   "86_Times_STEP_MAX_TIME_STP_010(1)" : Time = PLC "86_Times".STEP_MAX_TIME_STP_010 AT %DB1.DBW0, 1 s
   "86_Times_STEP_MAX_TIME_STP_020(1)" : Time = PLC "86_Times".STEP_MAX_TIME_STP_020 AT %DB1.DBW0, 1 s
   "86_Times_STEP_MAX_TIME_STP_030(1)" : Time = PLC "86_Times".STEP_MAX_TIME_STP_030 AT %DB1.DBW0, 1 s
   "86_Times_STEP_MAX_TIME_STP_040(1)" : Time = PLC "86_Times".STEP_MAX_TIME_STP_040 AT %DB1.DBW0, 1 s
   "86_Times_STEP_MAX_TIME_STP_050(1)" : Time = PLC "86_Times".STEP_MAX_TIME_STP_050 AT %DB1.DBW0, 1 s
   "86_Times_STEP_MAX_TIME_STP_060(1)" : Time = PLC "86_Times".STEP_MAX_TIME_STP_060 AT %DB1.DBW0, 1 s
   "86_Times_STEP_MAX_TIME_STP_070(1)" : Time = PLC "86_Times".STEP_MAX_TIME_STP_070 AT %DB1.DBW0, 1 s
   "86_Times_STEP_MAX_TIME_STP_080(1)" : Time = PLC "86_Times".STEP_MAX_TIME_STP_080 AT %DB1.DBW0, 1 s
   "86_Times_STEP_MAX_TIME_STP_090(1)" : Time = PLC "86_Times".STEP_MAX_TIME_STP_090 AT %DB1.DBW0, 1 s
   "86_Times_STEP_MAX_TIME_STP_100(1)" : Time = PLC "86_Times".STEP_MAX_TIME_STP_100 AT %DB1.DBW0, 1 s
   "86_Times_STEP_MAX_TIME_STP_110(1)" : Time = PLC "86_Times".STEP_MAX_TIME_STP_110 AT %DB1.DBW0, 1 s
   "86_Times_STEP_MAX_TIME_STP_120(1)" : Time = PLC "86_Times".STEP_MAX_TIME_STP_120 AT %DB1.DBW0, 1 s
   "86_Times_STEP_MAX_TIME_STP_130(1)" : Time = PLC "86_Times".STEP_MAX_TIME_STP_130 AT %DB1.DBW0, 1 s
   "86_Times_STEP_MAX_TIME_STP_140(1)" : Time = PLC "86_Times".STEP_MAX_TIME_STP_140 AT %DB1.DBW0, 1 s
   "86_Times_STEP_MAX_TIME_STP_150(1)" : Time = PLC "86_Times".STEP_MAX_TIME_STP_150 AT %DB1.DBW0, 1 s
   "86_Times_STEP_MAX_TIME_STP_160(1)" : Time = PLC "86_Times".STEP_MAX_TIME_STP_160 AT %DB1.DBW0, 1 s
   "86_Times_STEP_MAX_TIME_STP_170(1)" : Time = PLC "86_Times".STEP_MAX_TIME_STP_170 AT %DB1.DBW0, 1 s
   "86_Times_STEP_MAX_TIME_STP_180(1)" : Time = PLC "86_Times".STEP_MAX_TIME_STP_180 AT %DB1.DBW0, 1 s
   "86_Times_STEP_MAX_TIME_STP_190(1)" : Time = PLC "86_Times".STEP_MAX_TIME_STP_190 AT %DB1.DBW0, 1 s
   "86_Times_STEP_MAX_TIME_STP_200(1)" : Time = PLC "86_Times".STEP_MAX_TIME_STP_200 AT %DB1.DBW0, 1 s
   "86_Times_STEP_MAX_TIME_STP_210(1)" : Time = PLC "86_Times".STEP_MAX_TIME_STP_210 AT %DB1.DBW0, 1 s
   "86_Times_STEP_MAX_TIME_STP_220(1)" : Time = PLC "86_Times".STEP_MAX_TIME_STP_220 AT %DB1.DBW0, 1 s
   "86_Times_STEP_MAX_TIME_STP_230(1)" : Time = PLC "86_Times".STEP_MAX_TIME_STP_230 AT %DB1.DBW0, 1 s
   "86_Times_STEP_MAX_TIME_STP_240(1)" : Time = PLC "86_Times".STEP_MAX_TIME_STP_240 AT %DB1.DBW0, 1 s
   "86_Times_STEP_MAX_TIME_STP_250(1)" : Time = PLC "86_Times".STEP_MAX_TIME_STP_250 AT %DB1.DBW0, 1 s
   "86_Times_STEP_MAX_TIME_STP_260(1)" : Time = PLC "86_Times".STEP_MAX_TIME_STP_260 AT %DB1.DBW0, 1 s
   "86_Times_STEP_MAX_TIME_STP_270(1)" : Time = PLC "86_Times".STEP_MAX_TIME_STP_270 AT %DB1.DBW0, 1 s
   "86_Times_STEP_MAX_TIME_STP_280(1)" : Time = PLC "86_Times".STEP_MAX_TIME_STP_280 AT %DB1.DBW0, 1 s
   "86_Times_STEP_MAX_TIME_STP_290(1)" : Time = PLC "86_Times".STEP_MAX_TIME_STP_290 AT %DB1.DBW0, 1 s
   "86_Times_STEP_MAX_TIME_STP_300(1)" : Time = PLC "86_Times".STEP_MAX_TIME_STP_300 AT %DB1.DBW0, 1 s
   "86_Times_STEP_MAX_TIME_STP_310(1)" : Time = PLC "86_Times".STEP_MAX_TIME_STP_310 AT %DB1.DBW0, 1 s
   "86_Times_STEP_MAX_TIME_STP_320(1)" : Time = PLC "86_Times".STEP_MAX_TIME_STP_320 AT %DB1.DBW0, 1 s
   "86_Times_STEP_MAX_TIME_STP_330(1)" : Time = PLC "86_Times".STEP_MAX_TIME_STP_330 AT %DB1.DBW0, 1 s
   "86_Times_STEP_MAX_TIME_STP_340(1)" : Time = PLC "86_Times".STEP_MAX_TIME_STP_340 AT %DB1.DBW0, 1 s
   "86_Times_STEP_MAX_TIME_STP_350(1)" : Time = PLC Alarms_Acknowledge.IGG_ALARM_ACKNLG_2 AT %DB1.DBW0, 1 s
   "86_Times_STEP_MAX_TIME_STP_360(1)" : Time = PLC "86_Times".STEP_MAX_TIME_STP_360 AT %DB1.DBW0, 1 s
   "86_Times_STEP_MAX_TIME_STP_370(1)" : Time = PLC "86_Times".STEP_MAX_TIME_STP_370 AT %DB1.DBW0, 1 s
   "86_Times_STEP_MAX_TIME_STP_380(1)" : Time = PLC "86_Times".STEP_MAX_TIME_STP_380 AT %DB1.DBW0, 1 s
   "86_Times_STEP_MAX_TIME_STP_390(1)" : Time = PLC "86_Times".STEP_MAX_TIME_STP_390 AT %DB1.DBW0, 1 s
   "86_Times_STEP_MAX_TIME_STP_400(1)" : Time = PLC "86_Times".STEP_MAX_TIME_STP_400 AT %DB1.DBW0, 1 s
   "86_Times_STEP_MAX_TIME_STP_410(1)" : Time = PLC "86_Times".STEP_MAX_TIME_STP_410 AT %DB1.DBW0, 1 s
   "86_Times_STEP_MAX_TIME_STP_420(1)" : Time = PLC "86_Times".STEP_MAX_TIME_STP_420 AT %DB1.DBW0, 1 s
   "86_Times_STEP_MAX_TIME_STP_430(1)" : Time = PLC "86_Times".STEP_MAX_TIME_STP_430 AT %DB1.DBW0, 1 s
   "86_Times_STEP_MAX_TIME_STP_440(1)" : Time = PLC "86_Times".STEP_MAX_TIME_STP_440 AT %DB1.DBW0, 1 s
   "86_Times_STEP_MAX_TIME_STP_450(1)" : Time = PLC "86_Times".STEP_MAX_TIME_STP_450 AT %DB1.DBW0, 1 s
   "86_Times_STEP_MAX_TIME_STP_460(1)" : Time = PLC "86_Times".STEP_MAX_TIME_STP_460 AT %DB1.DBW0, 1 s
   "86_Times_STEP_MAX_TIME_STP_470(1)" : Time = PLC "86_Times".STEP_MAX_TIME_STP_470 AT %DB1.DBW0, 1 s
   "86_Times_STEP_MAX_TIME_STP_480(1)" : Time = PLC "86_Times".STEP_MAX_TIME_STP_480 AT %DB1.DBW0, 1 s
   "86_Times_STEP_MAX_TIME_STP_490(1)" : Time = PLC "86_Times".STEP_MAX_TIME_STP_490 AT %DB1.DBW0, 1 s
   "86_Times_STEP_MAX_TIME_STP_500(1)" : Time = PLC "86_Times".STEP_MAX_TIME_STP_500 AT %DB1.DBW0, 1 s
   "86_Times_STEP_MAX_TIME_STP_510(1)" : Time = PLC "86_Times".STEP_MAX_TIME_STP_510 AT %DB1.DBW0, 1 s
   "86_Times_STEP_MAX_TIME_STP_520(1)" : Time = PLC "86_Times".STEP_MAX_TIME_STP_520 AT %DB1.DBW0, 1 s
   "86_Times_STEP_MAX_TIME_STP_530(1)" : Time = PLC "86_Times".STEP_MAX_TIME_STP_530 AT %DB1.DBW0, 1 s
   "86_Times_STEP_MAX_TIME_STP_540(1)" : Time = PLC "86_Times".STEP_MAX_TIME_STP_540 AT %DB1.DBW0, 1 s
   "86_Times_STEP_MAX_TIME_STP_550(1)" : Time = PLC "86_Times".STEP_MAX_TIME_STP_550 AT %DB1.DBW0, 1 s
   "86_Times_STEP_MAX_TIME_STP_560(1)" : Time = PLC "86_Times".STEP_MAX_TIME_STP_560 AT %DB1.DBW0, 1 s
   "86_Times_STEP_MAX_TIME_STP_570(1)" : Time = PLC "10_DI_DATA".R3_SPR_DI_136_0 AT %DB1.DBW0, 1 s

HMI tags "IGG_HMI_Tags"
   "10_DI_Data_CV311_OPN" : Bool = PLC "10_DI_Data".CV311_OPN AT %DB1.DBW0, 1 s
   "10_DI_Data_CV311_CLSD" : Bool = PLC "82_To_HMI"."I&A Compressor Service Due" AT %DB1.DBW0, 1 s
   "80_From_HMI_RUN_IGG" : Bool = PLC "80_From_HMI".RUN_IGG AT %DB1.DBX0.0, 1 s
   "82_To_HMI_CA Blower Animation" : Int = PLC "82_To_HMI"."CA Blower Animation" AT %DB1.DBX0.0, 100 ms
   "10_DI_Data_E500B_ENBLD" : Bool = PLC "10_DI_Data".E500B_ENBLD AT %DB1.DBX0.0, 1 s
   "10_DI_Data_E500A_ENBLD" : Bool = PLC "10_DI_Data".E500A_ENBLD AT %DB1.DBX0.0, 1 s
   "80_From_HMI_RUN_IGG(1)" : Bool = PLC "80_From_HMI".RUN_IGG AT %DB1.DBX0.0, 1 s
   "14_DQ_Data_E500A_CNTRL" : Bool = PLC "14_DQ_Data".E500A_CNTRL AT %DB1.DBX0.0, 1 s
   "14_DQ_Data_E500B_CNTRL" : Bool = PLC "14_DQ_Data".E500B_CNTRL AT %DB1.DBX0.0, 1 s
   "82_To_HMI_Run Time A" : LTime = PLC "82_To_HMI"."Run Time A" AT %DB1.DBD0, 1 s
   "82_To_HMI_Run Time B" : LTime = PLC "82_To_HMI"."Run Time B" AT %DB1.DBD0, 1 s
   "80_From_HMI_SW_DTY_PMP_E500" : Bool = PLC "80_From_HMI".SW_DTY_PMP_E500 AT %DB1.DBW0, 1 s
   "12_AI_Data_PIT316_SCALED" : Real = PLC "12_AI_Data".PIT316_SCALED AT %DB1.DBX0.0, 1 s
   "12_AI_Data_TIT319_SCALED" : Real = PLC "12_AI_Data".TIT319_SCALED AT %DB1.DBX0.0, 1 s
   "12_AI_Data_TIT360_SCALED" : Real = PLC "12_AI_Data".TIT360_SCALED AT %DB1.DBX0.0, 1 s
   "12_AI_Data_PIT102_SCALED(1)" : Real = PLC "12_AI_Data".PIT102_SCALED AT %DB1.DBX0.0, 1 s
   "12_AI_Data_CV403_SCALED(1)" : Real = PLC "12_AI_Data".CV403_SCALED AT %DB1.DBX0.0, 1 s
   "12_AI_Data_E139_RPM_SCALED" : Real = PLC "12_AI_Data".E139_RPM_SCALED AT %DB1.DBX0.0, 1 s
   "12_AI_Data_E139_AMPS_SCALED" : Real = PLC "12_AI_Data".E139_AMPS_SCALED AT %DB1.DBX0.0, 1 s
   "12_AI_Data_PIT402_SCALED" : Real = PLC "12_AI_Data".PIT402_SCALED AT %DB1.DBX0.0, 1 s
   "10_DI_Data_E500B_TRIPPED" : Bool = PLC "10_DI_Data".E500B_TRIPPED AT %DB1.DBX0.0, 1 s
   "10_DI_Data_IGG_ESTOP_OK" : Bool = PLC "10_DI_Data".IGG_ESTOP_OK AT %DB1.DBX0.0, 1 s
   "10_DI_Data_E500A_TRIPPED" : Bool = PLC "10_DI_Data".E500A_TRIPPED AT %DB1.DBX0.0, 1 s
   "10_DI_Data_E500B_TRIPPED(1)" : Bool = PLC "10_DI_Data".E500B_TRIPPED AT %DB1.DBX0.0, 1 s
   "10_DI_Data_E500A_ENBLD(1)" : Bool = PLC "10_DI_Data".E500A_ENBLD AT %DB1.DBX0.0, 1 s
   "10_DI_Data_E500B_ENBLD(1)" : Bool = PLC "10_DI_Data".E500B_ENBLD AT %DB1.DBX0.0, 1 s
   "10_DI_Data_CV401_OPN" : Bool = PLC "10_DI_Data".CV401_OPN AT %DB1.DBX0.0, 1 s
   "10_DI_Data_CV401_CLSD" : Bool = PLC "10_DI_Data".CV401_CLSD AT %DB1.DBX0.0, 1 s
   "10_DI_Data_CV321_OPN" : Bool = PLC "10_DI_Data".CV321_OPN AT %DB1.DBX0.0, 1 s
   "10_DI_Data_CV321_CLSD" : Bool = PLC "10_DI_Data".CV321_CLSD AT %DB1.DBX0.0, 1 s
   "10_DI_Data_CV322_OPN" : Bool = PLC "10_DI_Data".CV322_OPN AT %DB1.DBX0.0, 1 s
   "10_DI_Data_CV322_CLSD" : Bool = PLC "10_DI_Data".CV322_CLSD AT %DB1.DBX0.0, 1 s
   "10_DI_Data_BC_PLC_PWR_OK" : Bool = PLC "10_DI_Data".BC_PLC_PWR_OK AT %DB1.DBX0.0, 1 s
   "10_DI_Data_IGG_VNT_PWR_OK" : Bool = PLC "10_DI_Data".IGG_VNT_PWR_OK AT %DB1.DBX0.0, 1 s
   "10_DI_Data_MCC_VNT_PWR_OK" : Bool = PLC "10_DI_Data".MCC_VNT_PWR_OK AT %DB1.DBX0.0, 1 s
   "10_DI_Data_7T1_PWR_OK" : Bool = PLC "10_DI_Data".7T1_PWR_OK AT %DB1.DBX0.0, 1 s
   "10_DI_Data_7T2_PWR_OK" : Bool = PLC "10_DI_Data".7T2_PWR_OK AT %DB1.DBX0.0, 1 s
   "10_DI_Data_7T3_PWR_OK" : Bool = PLC "10_DI_Data".7T3_PWR_OK AT %DB1.DBX0.0, 1 s
   "10_DI_Data_MAINTD_24VDC_PWR_OK" : Bool = PLC "10_DI_Data".MAINTD_24VDC_PWR_OK AT %DB1.DBX0.0, 1 s
   "10_DI_Data_SFTY_SYS_IL" : Bool = PLC "10_DI_Data".SFTY_SYS_IL AT %DB1.DBX0.0, 1 s
   "14_DQ_Data_CV311_312_CNTRL" : Bool = PLC "14_DQ_Data".CV311_312_CNTRL AT %DB1.DBX0.0, 1 s
   "14_DQ_Data_CV321_322_CNTRL" : Bool = PLC "14_DQ_Data".CV321_322_CNTRL AT %DB1.DBX0.0, 1 s
   "14_DQ_Data_CV401_CNTRL" : Bool = PLC "14_DQ_Data".CV401_CNTRL AT %DB1.DBX0.0, 1 s
   "51_SLAVE_STATUS_P301_ENBLD" : Bool = PLC "51_SLAVE_STATUS".P301_ENBLD AT %DB51.DBX14.3, 1 s
   "14_DQ_Data_24K2" : Bool = PLC "14_DQ_Data".24K2 AT %DB1.DBX0.0, 1 s
   "14_DQ_Data_24K3" : Bool = PLC "14_DQ_Data".24K3 AT %DB1.DBX0.0, 1 s
   "14_DQ_Data_24K4" : Bool = PLC "14_DQ_Data".24K4 AT %DB1.DBX0.0, 1 s
   "14_DQ_Data_24PF1" : Bool = PLC "14_DQ_Data".24PF1 AT %DB1.DBX0.0, 1 s
   "14_DQ_Data_24K3(2)" : Bool = PLC "14_DQ_Data".24K3 AT %DB1.DBX0.0, 1 s
   "14_DQ_Data_24PF3" : Bool = PLC "14_DQ_Data".24PF3 AT %DB1.DBX0.0, 1 s
   "14_DQ_Data_24PF4" : Bool = PLC "14_DQ_Data".24PF4 AT %DB1.DBX0.0, 100 ms
   "12_AI_Data_PIT102_SCALED" : Real = PLC "12_AI_Data".PIT102_SCALED AT %DB1.DBX0.0, 1 s
   "12_AI_Data_TIT401_SCALED" : Real = PLC "12_AI_Data".TIT401_SCALED AT %DB1.DBX0.0, 1 s
   "12_AI_Data_TIT315_SCALED" : Real = PLC "12_AI_Data".TIT315_SCALED AT %DB1.DBX0.0, 1 s
   "80_From_HMI_Request_Manual(1)" : Bool = PLC "80_From_HMI".Request_Manual AT %DB1.DBX0.0, 1 s
   "12_AI_Data_CV403_SCALED" : Real = PLC "12_AI_Data".CV403_SCALED AT %DB1.DBX0.0, 1 s
   "16_AQ_Data_CV403_CNTRL" : Real = PLC "16_AQ_Data".CV403_CNTRL AT %DB1.DBX0.0, 1 s
   "AlwaysTRUE" : Bool = PLC AlwaysTRUE AT %M1.2, 1 s
   "12_AI_Data_PIT359_SCALED" : Real = PLC "12_AI_Data".PIT359_SCALED AT %DB1.DBX0.0, 1 s
   "68_Sys_Status_Data_CSW_IL_PRES_IN_RNG" : Bool = PLC "68_Sys_Status_Data".CSW_IL_PRES_IN_RNG AT %DB1.DBX0.0, 1 s
   "14_DQ_Data_24PF2" : Bool = PLC "14_DQ_Data".24PF2 AT %DB1.DBX0.0, 1 s
   "19_AUTO_CMNDS_Data_PIT402_Target" : Real = PLC "19_AUTO_CMNDS_Data".PIT402_Target AT %DB1.DBD0, 1 s
   "80_From_HMI_RST_E500A_RT" : Bool = PLC "80_From_HMI".RST_E500A_RT AT %DB1.DBX0.0, 1 s
   "10_DI_Data_CV312_OPN" : Bool = PLC "10_DI_Data".CV312_OPN AT %DB1.DBX0.0, 1 s
   "10_DI_Data_CV312_CLSD" : Bool = PLC "10_DI_Data".CV312_CLSD AT %DB1.DBX0.0, 1 s
   "Clock_1Hz" : Bool = PLC Clock_1Hz AT %M0.5, 500 ms
   "14_DQ_Data_24K3(1)" : Bool = PLC "14_DQ_Data".24K3 AT %DB1.DBX0.0, 1 s
   "12_AI_Data_LIT305_SCALED" : Real = PLC "12_AI_Data".LIT305_SCALED AT %DB1.DBX0.0, 1 s
   "80_From_HMI_BWT_BYPASS(1)" : Bool = PLC "80_From_HMI".BWT_BYPASS AT %DB1.DBX0.0, 1 s
   "80_From_HMI_CRG_BLNK_MODE(1)" : Bool = PLC "80_From_HMI".CRG_BLNK_MODE AT %DB1.DBX0.0, 1 s
   "80_From_HMI_BWT_BYPASS" : Bool = PLC "80_From_HMI".BWT_BYPASS AT %DB1.DBX0.0, 1 s
   "80_From_HMI_CRG_BLNK_MODE" : Bool = PLC "80_From_HMI".CRG_BLNK_MODE AT %DB1.DBX0.0, 1 s
   "10_DI_Data_CV432_OPN" : Bool = PLC "10_DI_Data".CV432_OPN AT %DB1.DBX0.0, 1 s
   "10_DI_Data_CV432_CLSD" : Bool = PLC "10_DI_Data".CV432_CLSD AT %DB1.DBX0.0, 1 s
   "10_DI_Data_CV431_OPN" : Bool = PLC "10_DI_Data".CV431_OPN AT %DB1.DBX0.0, 1 s
   "10_DI_Data_CV431_CLSD" : Bool = PLC "10_DI_Data".CV431_CLSD AT %DB1.DBX0.0, 1 s
   "12_AI_Data_AT_O2_01_SCALED" : Real = PLC "12_AI_Data".AT_O2_01_SCALED AT %DB1.DBX0.0, 1 s
   "12_AI_Data_AT_O2_02_SCALED" : Real = PLC "12_AI_Data".AT_O2_02_SCALED AT %DB1.DBX0.0, 1 s
   "84_Setpoints_PIT102_Pilot_LowLow" : Real = PLC "84_Setpoints".PIT102_Pilot_LowLow AT %DB1.DBX0.0, 1 s
   "84_Setpoints_PIT102_Pilot_Low" : Real = PLC "84_Setpoints".PIT102_Pilot_Low AT %DB1.DBX0.0, 1 s
   "84_Setpoints_PIT102_Pilot_High" : Real = PLC "84_Setpoints".PIT102_Pilot_High AT %DB1.DBD0, 1 s
   "84_Setpoints_PIT102_Pilot_HighHigh" : Real = PLC "84_Setpoints".PIT102_Pilot_HighHigh AT %DB1.DBD0, 1 s
   "84_Setpoints_PIT102_Main_LowLow" : Real = PLC "84_Setpoints".PIT102_Main_LowLow AT %DB1.DBD0, 1 s
   "84_Setpoints_PIT102_Main_Low" : Real = PLC "84_Setpoints".PIT102_Main_Low AT %DB1.DBD0, 1 s
   "84_Setpoints_PIT102_Main_High" : Real = PLC "84_Setpoints".PIT102_Main_High AT %DB1.DBD0, 1 s
   "84_Setpoints_PIT102_Main_HighHigh" : Real = PLC "84_Setpoints".PIT102_Main_HighHigh AT %DB1.DBD0, 1 s
   "84_Setpoints_TIT401_High" : Real = PLC "84_Setpoints".TIT401_High AT %DB1.DBD0, 1 s
   "84_Setpoints_TIT401_HighHigh" : Real = PLC "84_Setpoints".TIT401_HighHigh AT %DB1.DBD0, 1 s
   "84_Setpoints_PIT402_Pilot_LowLow" : Real = PLC "84_Setpoints".PIT402_Pilot_LowLow AT %DB1.DBD0, 1 s
   "84_Setpoints_PIT402_Pilot_Low" : Real = PLC "84_Setpoints".PIT402_Pilot_Low AT %DB1.DBD0, 1 s
   "84_Setpoints_PIT402_Pilot_High" : Real = PLC "84_Setpoints".PIT402_Pilot_High AT %DB1.DBD0, 1 s
   "84_Setpoints_PIT402_Pilot_HighHigh" : Real = PLC "142_P304_HRS_RUN_DB".HRS AT %DB1.DBD0, 1 s
   "84_Setpoints_PIT402_Main_LowLow" : Real = PLC "84_Setpoints".PIT402_Main_LowLow AT %DB1.DBD0, 1 s
   "84_Setpoints_PIT402_Main_Low" : Real = PLC "84_Setpoints".PIT402_Main_Low AT %DB1.DBD0, 1 s
   "84_Setpoints_PIT402_Main_High" : Real = PLC "84_Setpoints".PIT402_Main_High AT %DB1.DBD0, 1 s
   "84_Setpoints_PIT402_Main_HighHigh" : Real = PLC "84_Setpoints".PIT402_Main_HighHigh AT %DB1.DBD0, 1 s
   "84_Setpoints_PIT112_LowLow" : Real = PLC "84_Setpoints".PIT112_LowLow AT %DB1.DBD0, 1 s
   "84_Setpoints_PIT112_Low" : Real = PLC "84_Setpoints".PIT112_Low AT %DB1.DBD0, 1 s
   "84_Setpoints_PIT112_High" : Real = PLC "84_Setpoints".PIT112_High AT %DB1.DBD0, 1 s
   "84_Setpoints_PIT112_HighHigh" : Real = PLC "84_Setpoints".PIT112_HighHigh AT %DB1.DBD0, 1 s
   "84_Setpoints_TIT315_High" : Real = PLC "84_Setpoints".TIT315_High AT %DB1.DBX0.0, 1 s
   "84_Setpoints_TIT315_HighHigh" : Real = PLC "84_Setpoints".TIT315_HighHigh AT %DB1.DBD0, 1 s
   "84_Setpoints_TIT319_High" : Real = PLC "84_Setpoints".TIT319_High AT %DB1.DBD0, 1 s
   "84_Setpoints_TIT319_HighHigh" : Real = PLC "84_Setpoints".TIT319_HighHigh AT %DB1.DBD0, 1 s
   "84_Setpoints_TIT360_High" : Real = PLC "84_Setpoints".TIT360_High AT %DB1.DBD0, 1 s
   "84_Setpoints_TIT360_HighHigh" : Real = PLC "84_Setpoints".TIT360_HighHigh AT %DB1.DBD0, 1 s
   "84_Setpoints_PIT359_LowLow" : Real = PLC "84_Setpoints".PIT359_LowLow AT %DB1.DBD0, 1 s
   "84_Setpoints_PIT359_Low" : Real = PLC "84_Setpoints".PIT359_Low AT %DB1.DBD0, 1 s
   "84_Setpoints_PIT359_High" : Real = PLC "84_Setpoints".PIT359_High AT %DB1.DBD0, 1 s
   "84_Setpoints_PIT359_HighHigh" : Real = PLC "84_Setpoints".PIT359_HighHigh AT %DB1.DBD0, 1 s
   "84_Setpoints_PIT316_LowLow" : Real = PLC "84_Setpoints".PIT316_LowLow AT %DB1.DBD0, 1 s
   "84_Setpoints_PIT316_Low" : Real = PLC "84_Setpoints".PIT316_Low AT %DB1.DBD0, 1 s
   "84_Setpoints_PIT316_High" : Real = PLC "84_Setpoints".PIT316_High AT %DB1.DBD0, 1 s
   "84_Setpoints_PIT316_HighHigh" : Real = PLC "84_Setpoints".PIT316_HighHigh AT %DB1.DBD0, 1 s
   "14_DQ_Data_CV431_432_CNTRL" : Bool = PLC "14_DQ_Data".CV431_432_CNTRL AT %DB1.DBX0.0, 1 s
   "14_DQ_Data_R2_SPR_DQ_0_7" : Bool = PLC "14_DQ_Data".R2_SPR_DQ_0_7 AT %DB1.DBX0.0, 1 s
   "14_DQ_Data_R2_SPR_DQ_1_0" : Bool = PLC "14_DQ_Data".R2_SPR_DQ_1_0 AT %DB1.DBX0.0, 1 s
   "80_From_HMI_MAN_DQ_0_0" : Bool = PLC "80_From_HMI".MAN_DQ_0_0 AT %DB1.DBX0.0, 1 s
   "80_From_HMI_MAN_DQ_0_1" : Bool = PLC "80_From_HMI".MAN_DQ_0_1 AT %DB1.DBX0.0, 1 s
   "80_From_HMI_MAN_DQ_0_2" : Bool = PLC "80_From_HMI".MAN_DQ_0_2 AT %DB1.DBX0.0, 1 s
   "80_From_HMI_MAN_DQ_0_3" : Bool = PLC "80_From_HMI".MAN_DQ_0_3 AT %DB1.DBX0.0, 1 s
   "80_From_HMI_MAN_DQ_0_4" : Bool = PLC "80_From_HMI".MAN_DQ_0_4 AT %DB1.DBX0.0, 1 s
   "80_From_HMI_MAN_DQ_0_5" : Bool = PLC "80_From_HMI".MAN_DQ_0_5 AT %DB1.DBX0.0, 1 s
   "80_From_HMI_MAN_DQ_0_6" : Bool = PLC "80_From_HMI".MAN_DQ_0_6 AT %DB1.DBX0.0, 1 s
   "80_From_HMI_MAN_DQ_0_7(1)" : Bool = PLC "80_From_HMI".MAN_DQ_0_7 AT %DB1.DBX0.0, 1 s
   "80_From_HMI_MAN_DQ_1_0(1)" : Bool = PLC "80_From_HMI".MAN_DQ_1_0 AT %DB1.DBX0.0, 1 s
   "80_From_HMI_MAN_DQ_1_1" : Bool = PLC "80_From_HMI".MAN_DQ_1_1 AT %DB1.DBX0.0, 1 s
   "80_From_HMI_MAN_DQ_1_2" : Bool = PLC "80_From_HMI".MAN_DQ_1_2 AT %DB1.DBX0.0, 1 s
   "80_From_HMI_MAN_DQ_1_3" : Bool = PLC "80_From_HMI".MAN_DQ_1_3 AT %DB1.DBX0.0, 1 s
   "80_From_HMI_MAN_DQ_1_4" : Bool = PLC "80_From_HMI".MAN_DQ_1_4 AT %DB1.DBX0.0, 1 s
   "80_From_HMI_MAN_DQ_1_5" : Bool = PLC "80_From_HMI".MAN_DQ_1_5 AT %DB1.DBX0.0, 1 s
   "80_From_HMI_MAN_DQ_1_6(1)" : Bool = PLC "80_From_HMI".MAN_DQ_1_6 AT %DB1.DBX0.0, 1 s
   "80_From_HMI_MAN_DQ_1_7" : Bool = PLC "80_From_HMI".MAN_DQ_1_7 AT %DB1.DBX0.0, 1 s
   "10_DI_Data_E139_READY" : Bool = PLC "10_DI_Data".E139_READY AT %DB1.DBX0.0, 1 s
   "10_DI_Data_E139_RUNNING(1)" : Bool = PLC "10_DI_Data".E139_RUNNING AT %DB1.DBX0.0, 1 s
   "10_DI_Data_E139_VSD_FLT" : Bool = PLC "10_DI_Data".E139_VSD_FLT AT %DB1.DBX0.0, 1 s
   "10_DI_Data_MCCP_5PG1_OK" : Bool = PLC "10_DI_Data".MCCP_5PG1_OK AT %DB1.DBX0.0, 1 s
   "10_DI_Data_R1_SPR_DI_3_7" : Bool = PLC "10_DI_Data".R1_SPR_DI_3_7 AT %DB1.DBX0.0, 1 s
   "84_Setpoints_AT_O2_1_Low" : Real = PLC "84_Setpoints".AT_O2_1_Low AT %DB1.DBD0, 1 s
   "84_Setpoints_PIT402_Main_Target" : Real = PLC "84_Setpoints".PIT402_Main_Target AT %DB1.DBX0.0, 1 s
   "84_Setpoints_PIT402_Pilot_Target" : Real = PLC "84_Setpoints".PIT402_Pilot_Target AT %DB1.DBD0, 1 s
   "14_DQ_Data_E139_CNTRL" : Bool = PLC RIO6_SPR_DI_63_7 AT %DB1.DBX0.0, 1 s
   "80_From_HMI_E139_SET_SPEED" : Real = PLC "80_From_HMI".E139_SET_SPEED AT %DB1.DBX0.0, 1 s
   "10_DI_Data_CV311_OPN(1)" : Bool = PLC "10_DI_Data".CV311_OPN AT %DB1.DBX0.0, 1 s
   "80_From_HMI_MAX_E500_RT" : LTime = PLC "80_From_HMI".MAX_E500_RT AT %DB1.DBX0.0, 1 s
   "68_Sys_Status_Data_IA_PRES_IN_RNG(1)" : Bool = PLC "68_Sys_Status_Data".IA_PRES_IN_RNG AT %DB1.DBX0.0, 1 s
   "68_Sys_Status_Data_FUEL_PRES_IN_RNG(1)" : Bool = PLC "68_Sys_Status_Data".FUEL_PRES_IN_RNG AT %DB1.DBX0.0, 1 s
   "16_AQ_Data_E139_SPEED" : Real = PLC "16_AQ_Data".E139_SPEED AT %DB1.DBD0, 1 s
   "16_AQ_Data_R1_SPR_AQ_102" : Real = PLC "16_AQ_Data".R1_SPR_AQ_102 AT %DB1.DBD0, 1 s
   "16_AQ_Data_R1_SPR_AQ_104" : Real = PLC "16_AQ_Data".R1_SPR_AQ_104 AT %DB1.DBD0, 1 s
   "80_From_HMI_MAN_AQ_INC_98(1)" : Bool = PLC "80_From_HMI".MAN_AQ_INC_98 AT %DB1.DBX0.0, 1 s
   "80_From_HMI_MAN_AQ_DEC_98(1)" : Bool = PLC "80_From_HMI".MAN_AQ_DEC_98 AT %DB1.DBX0.0, 1 s
   "80_From_HMI_MAN_AQ_INC_100" : Bool = PLC "80_From_HMI".MAN_AQ_INC_100 AT %DB1.DBX0.0, 1 s
   "80_From_HMI_MAN_AQ_DEC_100" : Bool = PLC "80_From_HMI".MAN_AQ_DEC_100 AT %DB1.DBX0.0, 1 s
   "80_From_HMI_MAN_AQ_INC_102(1)" : Bool = PLC "80_From_HMI".MAN_AQ_INC_102 AT %DB1.DBX0.0, 1 s
   "80_From_HMI_MAN_AQ_DEC_102(1)" : Bool = PLC "80_From_HMI".MAN_AQ_DEC_102 AT %DB1.DBX0.0, 1 s
   "80_From_HMI_MAN_AQ_DEC_104" : Bool = PLC "80_From_HMI".MAN_AQ_DEC_104 AT %DB1.DBX0.0, 1 s
   "80_From_HMI_MAN_AQ_INC_104" : Bool = PLC "80_From_HMI".MAN_AQ_INC_104 AT %DB1.DBX0.0, 1 s
   "80_From_HMI_STOP_IGG" : Bool = PLC "80_From_HMI".STOP_IGG AT %DB1.DBX0.0, 1 s
   "80_From_HMI_Request_Auto(1)" : Bool = PLC "80_From_HMI".Request_Auto AT %DB1.DBX0.0, 1 s
   "80_From_HMI_RST_AUT_SEQ(1)" : Bool = PLC "80_From_HMI".RST_AUT_SEQ AT %DB1.DBX0.0, 1 s
   "80_From_HMI_FAT_Mode" : Bool = PLC "80_From_HMI".FAT_Mode AT %DB1.DBX0.0, 1 s
   "80_From_HMI_IGG_STND_ALN" : Bool = PLC "80_From_HMI".IGG_STND_ALN AT %DB1.DBX0.0, 1 s
   "80_From_HMI_P301_PRSNT(1)" : Bool = PLC "80_From_HMI".P301_PRSNT AT %DB1.DBX0.0, 1 s
   "80_From_HMI_CV312_PRSNT" : Bool = PLC "80_From_HMI".CV312_PRSNT AT %DB1.DBX0.0, 1 s
   "80_From_HMI_CV431_PRSNT" : Bool = PLC "80_From_HMI".CV431_PRSNT AT %DB1.DBX0.0, 1 s
   "80_From_HMI_CV432_PRSNT" : Bool = PLC "80_From_HMI".CV432_PRSNT AT %DB1.DBX0.0, 1 s
   "80_From_HMI_SLNCE_BZR" : Bool = PLC "80_From_HMI".SLNCE_BZR AT %DB1.DBX0.0, 1 s
   "84_Setpoints_PIT102_Post_LowLow" : Real = PLC "84_Setpoints".PIT102_Post_LowLow AT %DB1.DBD0, 1 s
   "84_Setpoints_PIT102_Post_Low" : Real = PLC "84_Setpoints".PIT102_Post_Low AT %DB1.DBD0, 1 s
   "84_Setpoints_PIT102_Post_HighHigh" : Real = PLC "84_Setpoints".PIT102_Post_HighHigh AT %DB1.DBD0, 1 s
   "84_Setpoints_PIT102_Post_High" : Real = PLC "84_Setpoints".PIT102_Post_High AT %DB1.DBD0, 1 s
   "12_AI_Data_R1_SPR_AI_126_SCALED" : Real = PLC "12_AI_Data".R1_SPR_AI_126_SCALED AT %DB1.DBX0.0, 1 s
   "12_AI_Data_R1_SPR_AI_132_SCALED" : Real = PLC "12_AI_Data".R1_SPR_AI_132_SCALED AT %DB1.DBD0, 1 s
   "84_Setpoints_PIT402_Post_High" : Real = PLC "84_Setpoints".PIT402_Post_High AT %DB1.DBD0, 1 s
   "84_Setpoints_PIT402_Post_HighHigh" : Real = PLC "84_Setpoints".PIT402_Post_HighHigh AT %DB1.DBD0, 1 s
   "84_Setpoints_PIT402_Post_Low" : Real = PLC "84_Setpoints".PIT402_Post_Low AT %DB1.DBD0, 1 s
   "84_Setpoints_PIT402_Post_LowLow" : Real = PLC "84_Setpoints".PIT402_Post_LowLow AT %DB1.DBD0, 1 s
   "84_Setpoints_PIT402_Pilot_Target(1)" : Real = PLC "84_Setpoints".PIT402_Pilot_Target AT %DB1.DBD0, 1 s
   "84_Setpoints_PIT402_Main_Target(1)" : Real = PLC "84_Setpoints".PIT402_Main_Target AT %DB1.DBD0, 1 s
   "84_Setpoints_PIT402_Post_Target_Start" : Real = PLC "84_Setpoints".PIT402_Post_Target_Start AT %DB1.DBD0, 1 s
   "84_Setpoints_PIT401_Post_Target_Max" : Real = PLC "84_Setpoints".PIT401_Post_Target_Max AT %DB1.DBD0, 1 s
   "86_Times_PRE_BC_STRT_CMND_DLY" : Time = PLC "86_Times".PRE_BC_STRT_CMND_DLY AT %DB1.DBD0, 1 s
   "86_Times_PRE_CV203_CLS_CMND_DLY" : Time = PLC "86_Times".PRE_CV203_CLS_CMND_DLY AT %DB1.DBD0, 1 s
   "86_Times_POST_P301_STOP_DLY" : Time = PLC "86_Times".POST_P301_STOP_DLY AT %DB1.DBD0, 1 s
   "86_Times_POST_CV311_CLS_DLY" : Time = PLC "86_Times".POST_CV311_CLS_DLY AT %DB1.DBD0, 1 s
   "86_Times_POST_CV321_OPN_DLY" : Time = PLC "86_Times".POST_CV321_OPN_DLY AT %DB1.DBD0, 1 s
   "86_Times_CV311_MAX_TRVL_TIME" : Time = PLC "86_Times".CV311_MAX_TRVL_TIME AT %DB1.DBD0, 1 s
   "86_Times_CV312_MAX_TRVL_TIME" : Time = PLC "86_Times".CV312_MAX_TRVL_TIME AT %DB1.DBD0, 1 s
   "86_Times_CV321_MAX_TRVL_TIME" : Time = PLC "86_Times".CV321_MAX_TRVL_TIME AT %DB1.DBD0, 1 s
   "86_Times_CV322_MAX_TRVL_TIME" : Time = PLC "86_Times".CV322_MAX_TRVL_TIME AT %DB1.DBD0, 1 s
   "86_Times_CV401_MAX_TRVL_TIME" : Time = PLC "86_Times".CV401_MAX_TRVL_TIME AT %DB1.DBD0, 1 s
   "86_Times_CV431_MAX_TRVL_TIME" : Time = PLC "86_Times".CV431_MAX_TRVL_TIME AT %DB1.DBD0, 1 s
   "86_Times_CV432_MAX_TRVL_TIME" : Time = PLC "86_Times".CV432_MAX_TRVL_TIME AT %DB1.DBD0, 1 s
   "86_Times_STEP_MAX_TIME_STP_001(2)" : Time = PLC "86_Times".STEP_MAX_TIME_STP_001 AT %DB1.DBW0, 1 s
   "86_Times_STEP_MAX_TIME_STP_005(2)" : Time = PLC "86_Times".STEP_MAX_TIME_STP_005 AT %DB1.DBW0, 1 s
   "86_Times_STEP_MAX_TIME_STP_010(2)" : Time = PLC "86_Times".STEP_MAX_TIME_STP_010 AT %DB1.DBW0, 1 s
   "86_Times_STEP_MAX_TIME_STP_020(2)" : Time = PLC "86_Times".STEP_MAX_TIME_STP_020 AT %DB1.DBW0, 1 s
   "86_Times_STEP_MAX_TIME_STP_030(2)" : Time = PLC "86_Times".STEP_MAX_TIME_STP_030 AT %DB1.DBW0, 1 s
   "86_Times_STEP_MAX_TIME_STP_040(2)" : Time = PLC "86_Times".STEP_MAX_TIME_STP_040 AT %DB1.DBW0, 1 s
   "86_Times_STEP_MAX_TIME_STP_050(2)" : Time = PLC "86_Times".STEP_MAX_TIME_STP_050 AT %DB1.DBW0, 1 s
   "86_Times_STEP_MAX_TIME_STP_060(2)" : Time = PLC "86_Times".STEP_MAX_TIME_STP_060 AT %DB1.DBW0, 1 s
   "86_Times_STEP_MAX_TIME_STP_070(2)" : Time = PLC "86_Times".STEP_MAX_TIME_STP_070 AT %DB1.DBW0, 1 s
   "86_Times_STEP_MAX_TIME_STP_080(2)" : Time = PLC "86_Times".STEP_MAX_TIME_STP_080 AT %DB1.DBW0, 1 s
   "86_Times_STEP_MAX_TIME_STP_090(2)" : Time = PLC "86_Times".STEP_MAX_TIME_STP_090 AT %DB1.DBW0, 1 s
   "86_Times_STEP_MAX_TIME_STP_100(2)" : Time = PLC "86_Times".STEP_MAX_TIME_STP_100 AT %DB1.DBW0, 1 s
   "86_Times_STEP_MAX_TIME_STP_110(2)" : Time = PLC "86_Times".STEP_MAX_TIME_STP_110 AT %DB1.DBW0, 1 s
   "86_Times_STEP_MAX_TIME_STP_120(2)" : Time = PLC "86_Times".STEP_MAX_TIME_STP_120 AT %DB1.DBW0, 1 s
   "86_Times_STEP_MAX_TIME_STP_130(2)" : Time = PLC "86_Times".STEP_MAX_TIME_STP_130 AT %DB1.DBW0, 1 s
   "86_Times_STEP_MAX_TIME_STP_140(2)" : Time = PLC "86_Times".STEP_MAX_TIME_STP_140 AT %DB1.DBW0, 1 s
   "86_Times_STEP_MAX_TIME_STP_150(2)" : Time = PLC "86_Times".STEP_MAX_TIME_STP_150 AT %DB1.DBW0, 1 s
   "86_Times_STEP_MAX_TIME_STP_160(2)" : Time = PLC "86_Times".STEP_MAX_TIME_STP_160 AT %DB1.DBW0, 1 s
   "86_Times_STEP_MAX_TIME_STP_170(2)" : Time = PLC "86_Times".STEP_MAX_TIME_STP_170 AT %DB1.DBW0, 1 s
   "86_Times_STEP_MAX_TIME_STP_180(2)" : Time = PLC "86_Times".STEP_MAX_TIME_STP_180 AT %DB1.DBW0, 1 s
   "86_Times_STEP_MAX_TIME_STP_190(2)" : Time = PLC "86_Times".STEP_MAX_TIME_STP_190 AT %DB1.DBW0, 1 s
   "86_Times_STEP_MAX_TIME_STP_200(2)" : Time = PLC "86_Times".STEP_MAX_TIME_STP_200 AT %DB1.DBW0, 1 s
   "86_Times_STEP_MAX_TIME_STP_210(2)" : Time = PLC "86_Times".STEP_MAX_TIME_STP_210 AT %DB1.DBW0, 1 s
   "86_Times_STEP_MAX_TIME_STP_220(2)" : Time = PLC "86_Times".STEP_MAX_TIME_STP_220 AT %DB1.DBW0, 1 s
   "86_Times_STEP_MAX_TIME_STP_230(2)" : Time = PLC "86_Times".STEP_MAX_TIME_STP_230 AT %DB1.DBW0, 1 s
   "86_Times_STEP_MAX_TIME_STP_240(2)" : Time = PLC "86_Times".STEP_MAX_TIME_STP_240 AT %DB1.DBW0, 1 s
   "86_Times_STEP_MAX_TIME_STP_250(2)" : Time = PLC "86_Times".STEP_MAX_TIME_STP_250 AT %DB1.DBW0, 1 s
   "86_Times_STEP_MAX_TIME_STP_260(2)" : Time = PLC "86_Times".STEP_MAX_TIME_STP_260 AT %DB1.DBW0, 1 s
   "86_Times_STEP_MAX_TIME_STP_270(2)" : Time = PLC "86_Times".STEP_MAX_TIME_STP_270 AT %DB1.DBW0, 1 s
   "86_Times_STEP_MAX_TIME_STP_280(2)" : Time = PLC "86_Times".STEP_MAX_TIME_STP_280 AT %DB1.DBW0, 1 s
   "86_Times_STEP_MAX_TIME_STP_290(2)" : Time = PLC "86_Times".STEP_MAX_TIME_STP_290 AT %DB1.DBW0, 1 s
   "86_Times_STEP_MAX_TIME_STP_300(2)" : Time = PLC "86_Times".STEP_MAX_TIME_STP_300 AT %DB1.DBW0, 1 s
   "86_Times_STEP_MAX_TIME_STP_310(2)" : Time = PLC "86_Times".STEP_MAX_TIME_STP_310 AT %DB1.DBW0, 1 s
   "86_Times_STEP_MAX_TIME_STP_320(2)" : Time = PLC "86_Times".STEP_MAX_TIME_STP_320 AT %DB1.DBW0, 1 s
   "86_Times_STEP_MAX_TIME_STP_330(2)" : Time = PLC "86_Times".STEP_MAX_TIME_STP_330 AT %DB1.DBW0, 1 s
   "86_Times_STEP_MAX_TIME_STP_340(2)" : Time = PLC "86_Times".STEP_MAX_TIME_STP_340 AT %DB1.DBW0, 1 s
   "86_Times_STEP_MAX_TIME_STP_350(2)" : Time = PLC "86_Times".STEP_MAX_TIME_STP_350 AT %DB1.DBW0, 1 s
   "86_Times_STEP_MAX_TIME_STP_360(2)" : Time = PLC "86_Times".STEP_MAX_TIME_STP_360 AT %DB1.DBW0, 1 s
   "86_Times_STEP_MAX_TIME_STP_370(2)" : Time = PLC "86_Times".STEP_MAX_TIME_STP_370 AT %DB1.DBW0, 1 s
   "86_Times_STEP_MAX_TIME_STP_380(2)" : Time = PLC "86_Times".STEP_MAX_TIME_STP_380 AT %DB1.DBW0, 1 s
   "86_Times_STEP_MAX_TIME_STP_390(2)" : Time = PLC "86_Times".STEP_MAX_TIME_STP_390 AT %DB1.DBW0, 1 s
   "86_Times_STEP_MAX_TIME_STP_400(2)" : Time = PLC "86_Times".STEP_MAX_TIME_STP_400 AT %DB1.DBW0, 1 s
   "86_Times_STEP_MAX_TIME_STP_410(2)" : Time = PLC "86_Times".STEP_MAX_TIME_STP_410 AT %DB1.DBW0, 1 s
   "86_Times_STEP_MAX_TIME_STP_420(2)" : Time = PLC TT426_FPT_ALM_ANALOG_DB."LOW LEVEL VALUE (L)" AT %DB1.DBW0, 1 s
   "86_Times_STEP_MAX_TIME_STP_430(2)" : Time = PLC "86_Times".STEP_MAX_TIME_STP_430 AT %DB1.DBW0, 1 s
   "86_Times_STEP_MAX_TIME_STP_440(2)" : Time = PLC "86_Times".STEP_MAX_TIME_STP_440 AT %DB1.DBW0, 1 s
   "86_Times_STEP_MAX_TIME_STP_450(2)" : Time = PLC "86_Times".STEP_MAX_TIME_STP_450 AT %DB1.DBW0, 1 s
   "86_Times_STEP_MAX_TIME_STP_460(2)" : Time = PLC "86_Times".STEP_MAX_TIME_STP_460 AT %DB1.DBW0, 1 s
   "86_Times_STEP_MAX_TIME_STP_470(2)" : Time = PLC "86_Times".STEP_MAX_TIME_STP_470 AT %DB1.DBW0, 1 s
   "86_Times_STEP_MAX_TIME_STP_480(2)" : Time = PLC "86_Times".STEP_MAX_TIME_STP_480 AT %DB1.DBW0, 1 s
   "86_Times_STEP_MAX_TIME_STP_490(2)" : Time = PLC "86_Times".STEP_MAX_TIME_STP_490 AT %DB1.DBW0, 1 s
   "86_Times_STEP_MAX_TIME_STP_500(2)" : Time = PLC "86_Times".STEP_MAX_TIME_STP_500 AT %DB1.DBW0, 1 s
   "Logging SD Card Overflow" : Bool AT %DB1.DBX0.0
      on ChangeValue: "SD_Card_Overflow"()
   "88_treatment_POP_UP" : Bool = PLC "88_treatment".POP_UP AT %DB1.DBX0.0, 1 s
      on ChangeValue: "TreatmentdDailyChecks"()
   "88_treatment_POP_UP_CNFRM" : Bool = PLC "88_treatment".POP_UP_CNFRM AT %DB1.DBX0.0, 1 s

HMI tags "Warnings"
   "62_Warning_Data_BC_WARNING_WORD_01" : Word = PLC "62_Warning_Data".BC_WARNING_WORD_01 AT %DB62.DBW0, 1 s
   "62_Warning_Data_BC_WARNING_WORD_02" : Word = PLC "62_Warning_Data".BC_WARNING_WORD_02 AT %DB62.DBW2, 1 s
   "62_Warning_Data_BC_WARNING_WORD_03" : Word = PLC "62_Warning_Data".BC_WARNING_WORD_03 AT %DB62.DBW4, 1 s
   "62_Warning_Data_BC_WARNING_WORD_04" : Word = PLC "62_Warning_Data".BC_WARNING_WORD_04 AT %DB62.DBW6, 1 s
   "62_Warning_Data_BC_WARNING_WORD_05" : Word = PLC "62_Warning_Data".BC_WARNING_WORD_05 AT %DB62.DBW8, 1 s
   "62_Warning_Data_BC_WARNING_WORD_06" : Word = PLC "62_Warning_Data".BC_WARNING_WORD_06 AT %DB62.DBW10, 1 s
   "62_Warning_Data_GCU_WARNING_WORD_01" : Word = PLC "62_Warning_Data".GCU_WARNING_WORD_01 AT %DB62.DBW0, 1 s
   "62_Warning_Data_GCU_WARNING_WORD_02" : Word = PLC "62_Warning_Data".GCU_WARNING_WORD_02 AT %DB62.DBW2, 1 s
   "62_Warning_Data_GCU_WARNING_WORD_03" : Word = PLC "62_Warning_Data".GCU_WARNING_WORD_03 AT %DB62.DBW4, 1 s
   "62_Warning_Data_GCU_WARNING_WORD_04" : Word = PLC "62_Warning_Data".GCU_WARNING_WORD_04 AT %DB62.DBW6, 1 s
   "62_Warning_Data_GCU_WARNING_WORD_05" : Word = PLC "62_Warning_Data".GCU_WARNING_WORD_05 AT %DB62.DBW8, 1 s
   "62_Warning_Data_GCU_WARNING_WORD_06" : Word = PLC "62_Warning_Data".GCU_WARNING_WORD_06 AT %DB62.DBW10, 1 s
   "62_Warning_Data_GCU_WARNING_WORD_07" : Word = PLC "62_Warning_Data".GCU_WARNING_WORD_07 AT %DB62.DBW12, 1 s
   "62_Warning_Data_GCU_WARNING_WORD_08" : Word = PLC "62_Warning_Data".GCU_WARNING_WORD_08 AT %DB62.DBW14, 1 s
   "62_Warning_Data_GCU_WARNING_WORD_09" : Word = PLC "62_Warning_Data".GCU_WARNING_WORD_09 AT %DB62.DBW16, 1 s
   "62_Warning_Data_IGG_WARNING_WORD_01" : Word = PLC "62_Warning_Data".IGG_WARNING_WORD_01 AT %DB62.DBW0, 1 s
   "62_Warning_Data_IGG_WARNING_WORD_02" : Word = PLC "62_Warning_Data".IGG_WARNING_WORD_02 AT %DB62.DBW2, 1 s
   "62_Warning_Data_IGG_WARNING_WORD_03" : Word = PLC "62_Warning_Data".IGG_WARNING_WORD_03 AT %DB62.DBW4, 1 s
   "62_Warning_Data_IGG_WARNING_WORD_04" : Word = PLC "62_Warning_Data".IGG_WARNING_WORD_04 AT %DB62.DBW6, 1 s
   "62_Warning_Data_IGG_WARNING_WORD_05" : Word = PLC "62_Warning_Data".IGG_WARNING_WORD_05 AT %DB62.DBW8, 1 s
   "62_Warning_Data_IGG_WARNING_WORD_06" : Word = PLC "62_Warning_Data".IGG_WARNING_WORD_06 AT %DB62.DBW10, 1 s
   "2062_Warning_Data_BTCS_WARNING_WORD_01" : Word = PLC "2062_Warning_Data".BTCS_WARNING_WORD_01 AT %DB2062.DBW0, 1 s
   "2062_Warning_Data_BTCS_WARNING_WORD_02" : Word = PLC "2062_Warning_Data".BTCS_WARNING_WORD_02 AT %DB2062.DBW2, 1 s
   "2062_Warning_Data_BTCS_WARNING_WORD_03" : Word = PLC "2062_Warning_Data".BTCS_WARNING_WORD_03 AT %DB2062.DBW4, 1 s
   "2062_Warning_Data_BTCS_WARNING_WORD_04" : Word = PLC "2062_Warning_Data".BTCS_WARNING_WORD_04 AT %DB2062.DBW6, 1 s
   "2062_Warning_Data_BTCS_WARNING_WORD_05" : Word = PLC "2062_Warning_Data".BTCS_WARNING_WORD_05 AT %DB2062.DBW8, 1 s
   "2062_Warning_Data_BTCS_WARNING_WORD_06" : Word = PLC "2062_Warning_Data".BTCS_WARNING_WORD_06 AT %DB2062.DBW10, 1 s
   "2062_Warning_Data_BTCS_WARNING_WORD_07" : Word = PLC "2062_Warning_Data".BTCS_WARNING_WORD_07 AT %DB2062.DBW12, 1 s
   "2062_Warning_Data_BTCS_WARNING_WORD_08" : Word = PLC "2062_Warning_Data".BTCS_WARNING_WORD_08 AT %DB2062.DBW14, 1 s

